      ProcessValue <- "ST_Maintenance_g_u16_5_Times_TiShi_LongDai_Clean"
   Button "按钮_12" at 605,229 size 196x42; TextOff '1小时后提醒 / 1시간후 다시 알림'
      Visibility <- "ST_Maintenance_g_bo_5_Warn_Status_LongDai_Clean"
      on Click: ResetBit("ST_Maintenance_g_bo_5_Warn_Status_LongDai_Clean")
   Button "按钮_13" at 605,282 size 196x42; TextOff '已保养完毕 / 유지보수 이미 완료'; Authorization "User administration"
      Visibility <- "ST_Maintenance_g_bo_5_Warn_Status_LongDai_Clean"
      on Click: ResetBit("ST_Maintenance_g_bo_5_Status_LongDai_Clean")
   TextField "文本域_7" at 61,128 size 812x99; Text '保养时间到,请停机第 次为弓轴滚针 轴承加注黄油 保养时间到,请停机第 次为弓轴滚针 轴承加注黄油 유지보수시간. 기계 스톱. 제 차 보우축 니들 베어링에 그리스를 주입 한다.'
      Visibility <- "ST_Maintenance_g_bo_4_Warn_Status_GongZhou_Bearing"
   IOField "IO Field_90" at 368,129 size 70x28; FormatPattern 999
      Visibility <- "ST_Maintenance_g_bo_4_Warn_Status_GongZhou_Bearing"
      ProcessValue <- "ST_Maintenance_g_u16_4_Times_TiShi_GongZhou_Bearing"
   Button "按钮_10" at 628,129 size 196x42; TextOff '1小时后提醒 / 1시간후 다시 알림'
      Visibility <- "ST_Maintenance_g_bo_4_Warn_Status_GongZhou_Bearing"
      on Click: ResetBit("ST_Maintenance_g_bo_4_Warn_Status_GongZhou_Bearing")
   Button "按钮_11" at 628,182 size 196x42; TextOff '已保养完毕 / 유지보수 이미 완료'; Authorization "User administration"
      Visibility <- "ST_Maintenance_g_bo_4_Warn_Status_GongZhou_Bearing"
      on Click: ResetBit("ST_Maintenance_g_bo_4_Status_GongZhou_Bearing")
   TextField "文本域_9" at 42,238 size 812x100; Text '保养时间到,请停机第 次检查锭子传 动同步带:检查松紧度并适当调整 保养时间到,请停机第 次检查锭子传 动同步带:检查松紧度并适当调整 유지보수시간. 기계 스톱. 제 차 스핀들 전동 타이밍 벨트를 검사 : 조임 정도를 확인 하고 적당하게 조절한다.'
      Visibility <- "ST_Maintenance_g_bo_6_Warn_Status_DingZi_ChuanDong"
   IOField "IO Field_92" at 348,241 size 70x28; FormatPattern 999
      Visibility <- "ST_Maintenance_g_bo_6_Warn_Status_DingZi_ChuanDong"
      ProcessValue <- "ST_Maintenance_g_u16_6_Times_TiShi_DingZi_ChuanDong"
   Button "按钮_14" at 609,240 size 196x42; TextOff '1小时后提醒 / 1시간후 다시 알림'
      Visibility <- "ST_Maintenance_g_bo_6_Warn_Status_DingZi_ChuanDong"
      on Click: ResetBit("ST_Maintenance_g_bo_6_Warn_Status_DingZi_ChuanDong")
   Button "按钮_15" at 609,294 size 196x42; TextOff '已保养完毕 / 유지보수 이미 완료'; Authorization "User administration"
      Visibility <- "ST_Maintenance_g_bo_6_Warn_Status_DingZi_ChuanDong"
      on Click: ResetBit("ST_Maintenance_g_bo_6_Status_DingZi_ChuanDong")
   TextField "文本域_16" at 54,252 size 812x99; Text '保养时间到,请停机第 次清洁控制柜 卫生，用吸风机吸，注意不要用气管吹 保养时间到,请停机第 次清洁控制柜 卫生，用吸风机吸，注意不要用气管吹 유지보수시간. 기계 스톱. 제 차 제어함을 청소 하고 흡입팬으로 흡입한다. 주의할것은 에어 파이프로 불어서는 안된다.'
      Visibility <- "ST_Maintenance_g_bo_7_Warn_Status_ControlBox_Clean"
   IOField "IO Field_98" at 361,254 size 70x28; FormatPattern 999
      Visibility <- "ST_Maintenance_g_bo_7_Warn_Status_ControlBox_Clean"
      ProcessValue <- "ST_Maintenance_g_u16_7_Times_TiShi_ControlBox_Clean"
   Button "按钮_26" at 627,252 size 196x42; TextOff '1小时后提醒 / 1시간후 다시 알림'
      Visibility <- "ST_Maintenance_g_bo_7_Warn_Status_ControlBox_Clean"
      on Click: ResetBit("ST_Maintenance_g_bo_7_Warn_Status_ControlBox_Clean")
   Button "按钮_27" at 627,308 size 196x42; TextOff '已保养完毕 / 유지보수 이미 완료'; Authorization "User administration"
      Visibility <- "ST_Maintenance_g_bo_7_Warn_Status_ControlBox_Clean"
      on Click: ResetBit("ST_Maintenance_g_bo_7_Status_ControlBox_Clean")
   TextField "文本域_13" at 68,268 size 812x99; Text '保养时间到,请停机第 次清洁锭子电 机风扇上的绕毛 保养时间到,请停机第 次清洁锭子电 机风扇上的绕毛 유지보수시간. 기계 스톱. 제 차 스핀들 모터팬 에 감긴 원료 청소한다.'
      Visibility <- "ST_Maintenance_g_bo_8_Warn_Status_DingZi_Fan"
   IOField "IO Field_95" at 373,269 size 70x28; FormatPattern 999
      ProcessValue <- "ST_Maintenance_g_u16_8_Times_TiShi_DingZi_Fan"
      Visibility <- "ST_Maintenance_g_bo_8_Warn_Status_DingZi_Fan"
   Button "按钮_20" at 635,269 size 196x42; TextOff '1小时后提醒 / 1시간후 다시 알림'
      on Click: ResetBit("ST_Maintenance_g_bo_8_Warn_Status_DingZi_Fan")
      Visibility <- "ST_Maintenance_g_bo_8_Warn_Status_DingZi_Fan"
   Button "按钮_21" at 635,324 size 196x41; TextOff '已保养完毕 / 유지보수 이미 완료'; Authorization "User administration"
      on Click: ResetBit("ST_Maintenance_g_bo_8_Status_DingZi_Fan")
      Visibility <- "ST_Maintenance_g_bo_8_Warn_Status_DingZi_Fan"
   Button "按钮_6" at 742,567 size 137x44; TextOff '知道了 / OK'
      on Click: SetTag("ST_HMI_Var_HMI_i16_Dingzi_50102AlarmStatus", 0); ResetBit("ST_HMI_Var_HMI_bo_XiangLing")
      Visibility <- "ST_HMI_Var_HMI_i16_Dingzi_50102AlarmStatus"
   Circle "圆_1" at 782,478 size 60x60
      Visibility <- "ST_HMI_Var_HMI_i16_Dingzi_50102AlarmStatus"
      Appearance <- "ST_HMI_Var_HMI_bo_XiangLing"
   TextField "文本域_5" at 26,442 size 880x170; Text '锭子不转报警！请至报警画面解除报警，然后点击“退 出紧急停止”，点击“启动”开机，或者按正常步骤断电 重启，然后开机 스핀들이 돌아가지 않아 경보알림! 경보알림화면으로 이동하여 경보 해제후 "종료 비상 정지"를 클릭후 "시작"을 클릭하여 가동 하거나 정상적인 순서대로 단전 및 재부팅후 가동한다.'
      Visibility <- "ST_HMI_Var_HMI_i16_Dingzi_50102AlarmStatus"
   Button "按钮_16" at 751,544 size 137x44; TextOff '知道了 / OK'
      on Click: SetTag("ST_HMI_Var_HMI_i16_Dingzi_50102AlarmStatus", 0); ResetBit("ST_HMI_Var_HMI_bo_XiangLing")
      Visibility <- "ST_HMI_Var_HMI_i16_Dingzi_50102AlarmStatus"
   Circle "圆_3" at 791,455 size 60x60
      Visibility <- "ST_HMI_Var_HMI_i16_Dingzi_50102AlarmStatus"
      Appearance <- "ST_HMI_Var_HMI_bo_XiangLing"
   TextField "文本域_11" at 12,427 size 880x170; Text '捻度报警！设置捻度为 ， 实际捻度为 ， 已自动停止，请检查设置画面参数，重新设置总捻度， 检查设置其他参数，使画面上的参数没有红色闪烁，然 后按“启动”，若连续反复出现此报警，请从生头重新 开始 트위스트 경보 알림!설정 트위스트는 이고,실제 트위스트는 이며,이미 자동정지, 설정화면 매개변수를 확인하고,전체 트위스트를 다시 설정하고,기타 매개변수를 확인설정하여 화면의 매개변수에 빨간색이 깜 빡이지 않도록 해야 한다.그다음 "작동"을 누른다. 만약 이 경보가 연속 반 복적으로 나타나면 스레딩부터 다시 시작한다.'
      Visibility <- "ST_HMI_Var_HMI_i16_NianduAlarmStatus"
   IOField "IO Field_43" at 387,432 size 86x32; FormatPattern 9999
      on OnFinishInput: SetBit("ST_Calculation_Var_HMI_bo_Calculation_0_Start"); SetTag("ST_Calculation_Var_g_i16_Calculation_0_3_Select_Status", 1)
      Visibility <- "ST_HMI_Var_HMI_i16_NianduAlarmStatus"
      ProcessValue <- "ST_HMI_Var_HMI_r64NianDu_all"
   IOField "IO Field_3" at 691,432 size 86x32; FormatPattern 9999
      Visibility <- "ST_HMI_Var_HMI_i16_NianduAlarmStatus"
      ProcessValue <- "ST_HMI_Var_HMI_r64Niandu_all_Current"
   Button "按钮_7" at 745,537 size 137x44; TextOff '知道了 / OK'
      on Click: SetTag("ST_HMI_Var_HMI_i16_NianduAlarmStatus", 0); SetBit("ST_Calculation_Var_HMI_bo_Calculation_0_Start"); ResetBit("ST_HMI_Var_HMI_bo_XiangLing")
      Visibility <- "ST_HMI_Var_HMI_i16_NianduAlarmStatus"
   Circle "圆_2" at 785,448 size 60x60
      Visibility <- "ST_HMI_Var_HMI_i16_NianduAlarmStatus"
      Appearance <- "ST_HMI_Var_HMI_bo_XiangLing"

screen "动画" 1280x733, template "模板_2"
   on GenerateScreen: SetTag("变量_100", 9)
   Line "line_3" at 249,441 size 768x20
      Visibility <- "ST_HMI_Var_HMI_r64Axis_1_ZhangLi_Position_JuanRao_real2"
   Line "line_4" at 249,441 size 768x18
      Visibility <- "ST_HMI_Var_HMI_r64Axis_1_ZhangLi_Position_JuanRao_real2"
   Line "line_5" at 251,445 size 766x14
      Visibility <- "ST_HMI_Var_HMI_r64Axis_1_ZhangLi_Position_JuanRao_real2"
   Line "line_6" at 253,449 size 764x10
      Visibility <- "ST_HMI_Var_HMI_r64Axis_1_ZhangLi_Position_JuanRao_real2"
   Line "line_7" at 255,453 size 762x6
      Visibility <- "ST_HMI_Var_HMI_r64Axis_1_ZhangLi_Position_JuanRao_real2"
   Line "line_8" at 255,457 size 762x2
      Visibility <- "ST_HMI_Var_HMI_r64Axis_1_ZhangLi_Position_JuanRao_real2"
   Line "line_12" at 255,459 size 762x6
      Visibility <- "ST_HMI_Var_HMI_r64Axis_1_ZhangLi_Position_JuanRao_real2"
   Line "line_13" at 257,459 size 760x10
      Visibility <- "ST_HMI_Var_HMI_r64Axis_1_ZhangLi_Position_JuanRao_real2"
   Line "line_14" at 257,459 size 760x14
      Visibility <- "ST_HMI_Var_HMI_r64Axis_1_ZhangLi_Position_JuanRao_real2"
   Line "line_27" at 214,457 size 806x20
      Visibility <- "ST_HMI_Var_HMI_r64Axis_1_ZhangLi_Position_JuanRao_real2"
   Line "line_1" at 214,457 size 804x20
      Visibility <- "ST_Main_Var_g_i16_Automatic_Status"
   Group "Group_8" at 262,551 size 1011x176
   Bar "棒图_1" at 177,50 size 20x295; Unit r/min; MinimumValue 0; MaximumValue 10000
      ProcessValue <- "ST_HMI_Var_HMI_r64Axis_DingZi_Velocity_real"
   IOField "IO Field_57" at 166,346 size 62x30; FormatPattern 99999
      ProcessValue <- "ST_HMI_Var_HMI_r64Axis_DingZi_Velocity_real"
   Button "HmiScreenItemData_1" at 1115,95 size 159x60; TextOn '向后 / 後向き / 뒤로'; TextOff '向后 / 後向き / 뒤로'
      on Release: function_efd93a16()
   Rectangle "矩形_3" at 282,425 size 220x80
      DirectMovement <- "ST_HMI_Var_HMI_r64Axis_ZouChe_Position_real2"
   Rectangle "矩形_5" at 486,425 size 214x80
      DirectMovement <- "ST_HMI_Var_HMI_r64Axis_ZouChe_Position_real2"
   Rectangle "矩形_7" at 700,425 size 214x80
      DirectMovement <- "ST_HMI_Var_HMI_r64Axis_ZouChe_Position_real2"
   Rectangle "矩形_8" at 914,425 size 214x80
      DirectMovement <- "ST_HMI_Var_HMI_r64Axis_ZouChe_Position_real2"
   Group "Group_1" at 160,442 size 88x240
   Group "Group_2" at 20,9 size 90x480
   Group "Group_5" at 48,441 size 200x252
   Polyline "折线_1" at 163,442 size 85x231
      Visibility <- "ST_HMI_Var_HMI_r64Axis_ChengXing_Position_real2"
   Polyline "折线_25" at 179,442 size 69x179
      Visibility <- "ST_HMI_Var_HMI_r64Axis_ChengXing_Position_real2"
   Polyline "折线_37" at 197,442 size 51x118
      Visibility <- "ST_HMI_Var_HMI_r64Axis_ChengXing_Position_real2"
   Polyline "折线_45" at 213,442 size 35x57
      Visibility <- "ST_HMI_Var_HMI_r64Axis_ChengXing_Position_real2"
   Polyline "折线_46" at 169,442 size 79x233
      Visibility <- "ST_HMI_Var_HMI_r64Axis_ChengXing_Position_real2"
   Polyline "折线_50" at 179,442 size 69x181
      Visibility <- "ST_HMI_Var_HMI_r64Axis_ChengXing_Position_real2"
   Polyline "折线_51" at 197,442 size 51x122
      Visibility <- "ST_HMI_Var_HMI_r64Axis_ChengXing_Position_real2"
   Polyline "折线_57" at 213,442 size 35x60
      Visibility <- "ST_HMI_Var_HMI_r64Axis_ChengXing_Position_real2"
   Polyline "折线_68" at 169,442 size 79x235
      Visibility <- "ST_HMI_Var_HMI_r64Axis_ChengXing_Position_real2"
   Polyline "折线_71" at 179,442 size 69x184
      Visibility <- "ST_HMI_Var_HMI_r64Axis_ChengXing_Position_real2"
   Polyline "折线_72" at 197,442 size 51x124
      Visibility <- "ST_HMI_Var_HMI_r64Axis_ChengXing_Position_real2"
   Polyline "折线_77" at 213,442 size 35x63
      Visibility <- "ST_HMI_Var_HMI_r64Axis_ChengXing_Position_real2"
   Polyline "折线_78" at 163,442 size 85x237
      Visibility <- "ST_HMI_Var_HMI_r64Axis_ChengXing_Position_real2"
   Polyline "折线_79" at 175,442 size 73x187
      Visibility <- "ST_HMI_Var_HMI_r64Axis_ChengXing_Position_real2"
   Polyline "折线_80" at 191,442 size 57x127
      Visibility <- "ST_HMI_Var_HMI_r64Axis_ChengXing_Position_real2"
   Polyline "折线_81" at 207,442 size 41x66
      Visibility <- "ST_HMI_Var_HMI_r64Axis_ChengXing_Position_real2"
   Polyline "折线_82" at 160,442 size 88x240
      Visibility <- "ST_HMI_Var_HMI_r64Axis_ChengXing_Position_real2"
   Polyline "折线_83" at 207,442 size 41x69
      Visibility <- "ST_HMI_Var_HMI_r64Axis_ChengXing_Position_real2"
   Polyline "折线_84" at 197,442 size 51x131
      Visibility <- "ST_HMI_Var_HMI_r64Axis_ChengXing_Position_real2"
   Polyline "折线_85" at 175,442 size 73x190
      Visibility <- "ST_HMI_Var_HMI_r64Axis_ChengXing_Position_real2"
   Polyline "折线_86" at 175,442 size 73x192
      Visibility <- "ST_HMI_Var_HMI_r64Axis_ChengXing_Position_real2"
   Polyline "折线_87" at 187,442 size 61x133
      Visibility <- "ST_HMI_Var_HMI_r64Axis_ChengXing_Position_real2"
   Polyline "折线_88" at 207,442 size 41x72
      Visibility <- "ST_HMI_Var_HMI_r64Axis_ChengXing_Position_real2"
   Polyline "折线_89" at 179,442 size 69x195
      Visibility <- "ST_HMI_Var_HMI_r64Axis_ChengXing_Position_real2"
   Polyline "折线_90" at 185,442 size 63x136
      Visibility <- "ST_HMI_Var_HMI_r64Axis_ChengXing_Position_real2"
   Polyline "折线_91" at 207,442 size 41x75
      Visibility <- "ST_HMI_Var_HMI_r64Axis_ChengXing_Position_real2"
   Polyline "折线_92" at 175,442 size 73x198
      Visibility <- "ST_HMI_Var_HMI_r64Axis_ChengXing_Position_real2"
   Polyline "折线_93" at 191,442 size 57x140
      Visibility <- "ST_HMI_Var_HMI_r64Axis_ChengXing_Position_real2"
   Polyline "折线_94" at 207,442 size 41x78
      Visibility <- "ST_HMI_Var_HMI_r64Axis_ChengXing_Position_real2"
   Polyline "折线_95" at 175,442 size 73x199
      Visibility <- "ST_HMI_Var_HMI_r64Axis_ChengXing_Position_real2"
   Polyline "折线_96" at 185,442 size 63x143
      Visibility <- "ST_HMI_Var_HMI_r64Axis_ChengXing_Position_real2"
   Polyline "折线_97" at 201,442 size 47x81
      Visibility <- "ST_HMI_Var_HMI_r64Axis_ChengXing_Position_real2"
   Polyline "折线_98" at 175,442 size 73x202
      Visibility <- "ST_HMI_Var_HMI_r64Axis_ChengXing_Position_real2"
   Polyline "折线_99" at 191,442 size 57x146
      Visibility <- "ST_HMI_Var_HMI_r64Axis_ChengXing_Position_real2"
   Polyline "折线_100" at 207,442 size 41x84
      Visibility <- "ST_HMI_Var_HMI_r64Axis_ChengXing_Position_real2"
   Polyline "折线_101" at 167,442 size 81x205
      Visibility <- "ST_HMI_Var_HMI_r64Axis_ChengXing_Position_real2"
   Polyline "折线_102" at 185,442 size 63x149
      Visibility <- "ST_HMI_Var_HMI_r64Axis_ChengXing_Position_real2"
   Polyline "折线_103" at 201,442 size 47x87
      Visibility <- "ST_HMI_Var_HMI_r64Axis_ChengXing_Position_real2"
   Polyline "折线_104" at 169,442 size 79x207
      Visibility <- "ST_HMI_Var_HMI_r64Axis_ChengXing_Position_real2"
   Polyline "折线_105" at 201,442 size 47x91
      Visibility <- "ST_HMI_Var_HMI_r64Axis_ChengXing_Position_real2"
   Polyline "折线_106" at 191,442 size 57x153
      Visibility <- "ST_HMI_Var_HMI_r64Axis_ChengXing_Position_real2"
   Polyline "折线_107" at 169,442 size 79x211
      Visibility <- "ST_HMI_Var_HMI_r64Axis_ChengXing_Position_real2"
   Polyline "折线_108" at 185,442 size 63x156
      Visibility <- "ST_HMI_Var_HMI_r64Axis_ChengXing_Position_real2"
   Polyline "折线_109" at 201,442 size 47x94
      Visibility <- "ST_HMI_Var_HMI_r64Axis_ChengXing_Position_real2"
   Polyline "折线_110" at 169,442 size 79x213
      Visibility <- "ST_HMI_Var_HMI_r64Axis_ChengXing_Position_real2"
   Polyline "折线_111" at 201,442 size 47x96
      Visibility <- "ST_HMI_Var_HMI_r64Axis_ChengXing_Position_real2"
   Polyline "折线_112" at 185,442 size 63x159
      Visibility <- "ST_HMI_Var_HMI_r64Axis_ChengXing_Position_real2"
   Polyline "折线_113" at 170,442 size 78x216
      Visibility <- "ST_HMI_Var_HMI_r64Axis_ChengXing_Position_real2"
   Polyline "折线_114" at 185,442 size 63x161
      Visibility <- "ST_HMI_Var_HMI_r64Axis_ChengXing_Position_real2"
   Polyline "折线_115" at 201,442 size 47x100
      Visibility <- "ST_HMI_Var_HMI_r64Axis_ChengXing_Position_real2"
   Polyline "折线_116" at 179,442 size 69x165
      Visibility <- "ST_HMI_Var_HMI_r64Axis_ChengXing_Position_real2"
   Polyline "折线_117" at 169,442 size 79x219
      Visibility <- "ST_HMI_Var_HMI_r64Axis_ChengXing_Position_real2"
   Polyline "折线_118" at 201,442 size 47x104
      Visibility <- "ST_HMI_Var_HMI_r64Axis_ChengXing_Position_real2"
   Polyline "折线_119" at 169,442 size 79x221
      Visibility <- "ST_HMI_Var_HMI_r64Axis_ChengXing_Position_real2"
   Polyline "折线_120" at 201,442 size 47x106
      Visibility <- "ST_HMI_Var_HMI_r64Axis_ChengXing_Position_real2"
   Polyline "折线_121" at 185,442 size 63x168
      Visibility <- "ST_HMI_Var_HMI_r64Axis_ChengXing_Position_real2"
   Polyline "折线_122" at 169,442 size 79x223
      Visibility <- "ST_HMI_Var_HMI_r64Axis_ChengXing_Position_real2"
   Polyline "折线_123" at 179,442 size 69x170
      Visibility <- "ST_HMI_Var_HMI_r64Axis_ChengXing_Position_real2"
   Polyline "折线_124" at 197,442 size 51x109
      Visibility <- "ST_HMI_Var_HMI_r64Axis_ChengXing_Position_real2"
   Polyline "折线_125" at 165,442 size 83x225
      Visibility <- "ST_HMI_Var_HMI_r64Axis_ChengXing_Position_real2"
   Polyline "折线_126" at 193,442 size 55x112
      Visibility <- "ST_HMI_Var_HMI_r64Axis_ChengXing_Position_real2"
   Polyline "折线_127" at 179,442 size 69x173
      Visibility <- "ST_HMI_Var_HMI_r64Axis_ChengXing_Position_real2"
   Polyline "折线_128" at 169,442 size 79x228
      Visibility <- "ST_HMI_Var_HMI_r64Axis_ChengXing_Position_real2"
   Polyline "折线_129" at 197,442 size 51x115
      Visibility <- "ST_HMI_Var_HMI_r64Axis_ChengXing_Position_real2"
   Polyline "折线_130" at 179,442 size 69x176
      Visibility <- "ST_HMI_Var_HMI_r64Axis_ChengXing_Position_real2"
   Polygon "多边形_195" at 20,131 size 90x323
      Visibility <- "VBS_hengsi_status1"
   Polygon "多边形_196" at 20,229 size 90x225
      Visibility <- "VBS_hengsi_status1"
   Polygon "多边形_264" at 44,338 size 44x116
      Visibility <- "VBS_hengsi_status0"
   Polygon "多边形_265" at 49,350 size 34x104
      Visibility <- "VBS_hengsi_status0"
   Polygon "多边形_198" at 20,124 size 90x330
      Visibility <- "VBS_hengsi_status1"
   Polygon "多边形_199" at 20,223 size 90x231
      Visibility <- "VBS_hengsi_status1"
   Polygon "多边形_266" at 41,329 size 49x124
      Visibility <- "VBS_hengsi_status0"
   Polygon "多边形_201" at 20,120 size 90x334
      Visibility <- "VBS_hengsi_status1"
   Polygon "多边形_202" at 20,219 size 90x235
      Visibility <- "VBS_hengsi_status1"
   Polygon "多边形_267" at 38,319 size 54x135
      Visibility <- "VBS_hengsi_status0"
   Polygon "多边形_204" at 20,117 size 90x337
      Visibility <- "VBS_hengsi_status1"
   Polygon "多边形_205" at 20,213 size 90x241
      Visibility <- "VBS_hengsi_status1"
   Polygon "多边形_268" at 36,311 size 58x143
      Visibility <- "VBS_hengsi_status0"
   Polygon "多边形_207" at 20,113 size 90x341
      Visibility <- "VBS_hengsi_status1"
   Polygon "多边形_208" at 20,210 size 90x243
      Visibility <- "VBS_hengsi_status1"
   Polygon "多边形_269" at 35,306 size 60x148
      Visibility <- "VBS_hengsi_status0"
   Polygon "多边形_210" at 20,107 size 90x347
      Visibility <- "VBS_hengsi_status0"
   Polygon "多边形_211" at 20,206 size 90x248
      Visibility <- "VBS_hengsi_status1"
   Polygon "多边形_270" at 35,298 size 60x156
      Visibility <- "VBS_hengsi_status0"
   Polygon "多边形_213" at 20,103 size 90x351
      Visibility <- "VBS_hengsi_status1"
   Polygon "多边形_214" at 20,202 size 90x252
      Visibility <- "VBS_hengsi_status1"
   Polygon "多边形_271" at 34,292 size 63x162
      Visibility <- "VBS_hengsi_status0"
   Polygon "多边形_216" at 20,97 size 90x357
      Visibility <- "VBS_hengsi_status1"
   Polygon "多边形_217" at 20,196 size 90x258
      Visibility <- "VBS_hengsi_status1"
   Polygon "多边形_272" at 34,288 size 63x166
      Visibility <- "VBS_hengsi_status0"
   Polygon "多边形_219" at 20,93 size 90x361
      Visibility <- "VBS_hengsi_status1"
   Polygon "多边形_220" at 20,192 size 90x262
      Visibility <- "VBS_hengsi_status1"
   Polygon "多边形_273" at 32,285 size 66x169
      Visibility <- "VBS_hengsi_status0"
   Polygon "多边形_222" at 20,90 size 90x364
      Visibility <- "VBS_hengsi_status1"
   Polygon "多边形_223" at 20,189 size 90x265
      Visibility <- "VBS_hengsi_status1"
   Polygon "多边形_274" at 32,283 size 66x171
      Visibility <- "VBS_hengsi_status0"
   Polygon "多边形_225" at 20,86 size 90x368
      Visibility <- "VBS_hengsi_status1"
   Polygon "多边形_226" at 20,185 size 90x269
      Visibility <- "VBS_hengsi_status1"
   Polygon "多边形_275" at 31,279 size 68x175
      Visibility <- "VBS_hengsi_status0"
   Polygon "多边形_228" at 20,80 size 90x374
      Visibility <- "VBS_hengsi_status1"
   Polygon "多边形_229" at 20,179 size 90x275
      Visibility <- "VBS_hengsi_status1"
   Polygon "多边形_276" at 31,275 size 68x179
      Visibility <- "VBS_hengsi_status0"
   Polygon "多边形_231" at 20,76 size 90x378
      Visibility <- "VBS_hengsi_status1"
   Polygon "多边形_232" at 20,175 size 90x279
      Visibility <- "VBS_hengsi_status1"
   Polygon "多边形_277" at 29,271 size 70x183
      Visibility <- "VBS_hengsi_status0"
   Polygon "多边形_234" at 20,70 size 90x384
      Visibility <- "VBS_hengsi_status1"
   Polygon "多边形_235" at 20,169 size 90x285
      Visibility <- "VBS_hengsi_status1"
   Polygon "多边形_278" at 27,271 size 74x183
      Visibility <- "VBS_hengsi_status0"
   Polygon "多边形_237" at 20,69 size 90x385
      Visibility <- "VBS_hengsi_status1"
   Polygon "多边形_238" at 20,165 size 90x289
      Visibility <- "VBS_hengsi_status1"
   Polygon "多边形_279" at 27,267 size 74x187
      Visibility <- "VBS_hengsi_status0"
   Polygon "多边形_240" at 20,63 size 90x391
      Visibility <- "VBS_hengsi_status1"
   Polygon "多边形_241" at 20,162 size 90x292
      Visibility <- "VBS_hengsi_status1"
   Polygon "多边形_280" at 26,263 size 77x191
      Visibility <- "VBS_hengsi_status0"
   Polygon "多边形_243" at 20,59 size 90x395
      Visibility <- "VBS_hengsi_status1"
   Polygon "多边形_244" at 20,158 size 90x296
      Visibility <- "VBS_hengsi_status1"
   Polygon "多边形_281" at 26,261 size 77x193
      Visibility <- "VBS_hengsi_status0"
   Polygon "多边形_246" at 20,53 size 90x401
      Visibility <- "VBS_hengsi_status1"
   Polygon "多边形_247" at 20,152 size 90x302
      Visibility <- "VBS_hengsi_status1"
   Polygon "多边形_282" at 25,258 size 79x196
      Visibility <- "VBS_hengsi_status0"
   Polygon "多边形_249" at 20,49 size 90x405
      Visibility <- "VBS_hengsi_status1"
   Polygon "多边形_250" at 20,148 size 90x306
      Visibility <- "VBS_hengsi_status1"
   Polygon "多边形_283" at 25,254 size 79x200
      Visibility <- "VBS_hengsi_status0"
   Polygon "多边形_252" at 20,45 size 90x409
      Visibility <- "VBS_hengsi_status1"
   Polygon "多边形_253" at 20,142 size 90x312
      Visibility <- "VBS_hengsi_status1"
   Polygon "多边形_284" at 23,250 size 83x204
      Visibility <- "VBS_hengsi_status0"
   Polygon "多边形_255" at 20,42 size 90x412
      Visibility <- "VBS_hengsi_status1"
   Polygon "多边形_256" at 20,141 size 90x313
      Visibility <- "VBS_hengsi_status1"
   Polygon "多边形_285" at 23,246 size 83x208
      Visibility <- "VBS_hengsi_status0"
   Polygon "多边形_258" at 20,135 size 90x319
      Visibility <- "VBS_hengsi_status1"
   Polygon "多边形_286" at 22,242 size 85x212
      Visibility <- "VBS_hengsi_status0"
   Polygon "多边形_287" at 22,238 size 85x216
      Visibility <- "VBS_hengsi_status0"
   Polygon "多边形_288" at 20,237 size 88x217
      Visibility <- "VBS_hengsi_status0"
   Polygon "多边形_289" at 20,231 size 90x223
      Visibility <- "VBS_hengsi_status0"
   Group "Group_3" at 48,441 size 200x252
   Group "Group_4" at 48,441 size 200x252
   Line "线_1" at 68,549 size 180x9
      Visibility <- "ST_HMI_Var_HMI_r64Axis_ChengXing_Position_real2"
   Line "线_2" at 68,549 size 166x68
      Visibility <- "ST_HMI_Var_HMI_r64Axis_ChengXing_Position_real2"
   Line "线_136#mig1_2" at 68,549 size 132x120
      Visibility <- "ST_HMI_Var_HMI_r64Axis_ChengXing_Position_real2"
   Line "线_3" at 68,443 size 144x106
      Visibility <- "ST_HMI_Var_HMI_r64Axis_ChengXing_Position_real2"
   Line "线_4" at 68,497 size 172x52
      Visibility <- "ST_HMI_Var_HMI_r64Axis_ChengXing_Position_real2"
   Line "线_11#mig1_2" at 68,441 size 143x108
      Visibility <- "ST_HMI_Var_HMI_r64Axis_ChengXing_Position_real2"
   Line "线_5" at 68,501 size 173x48
      Visibility <- "ST_HMI_Var_HMI_r64Axis_ChengXing_Position_real2"
   Line "线_6" at 68,549 size 129x122
      Visibility <- "ST_HMI_Var_HMI_r64Axis_ChengXing_Position_real2"
   Line "线_157" at 68,446 size 146x103
      Visibility <- "ST_HMI_Var_HMI_r64Axis_ChengXing_Position_real2"
   Line "线_115#mig1_2" at 68,549 size 179x13
      Visibility <- "ST_HMI_Var_HMI_r64Axis_ChengXing_Position_real2"
   Line "线_7" at 68,549 size 165x71
      Visibility <- "ST_HMI_Var_HMI_r64Axis_ChengXing_Position_real2"
   Line "线_159" at 68,549 size 179x15
      Visibility <- "ST_HMI_Var_HMI_r64Axis_ChengXing_Position_real2"
   Line "线_8" at 68,549 size 163x74
      Visibility <- "ST_HMI_Var_HMI_r64Axis_ChengXing_Position_real2"
   Line "线_9" at 68,549 size 127x124
      Visibility <- "ST_HMI_Var_HMI_r64Axis_ChengXing_Position_real2"
   Line "线_13#mig1_2" at 68,448 size 147x101
      Visibility <- "ST_HMI_Var_HMI_r64Axis_ChengXing_Position_real2"
   Line "线_14" at 68,503 size 174x46
      Visibility <- "ST_HMI_Var_HMI_r64Axis_ChengXing_Position_real2"
   Line "线_22" at 68,549 size 179x18
      Visibility <- "ST_HMI_Var_HMI_r64Axis_ChengXing_Position_real2"
   Line "线_24" at 68,549 size 162x77
      Visibility <- "ST_HMI_Var_HMI_r64Axis_ChengXing_Position_real2"
   Line "线_25" at 68,549 size 125x126
      Visibility <- "ST_HMI_Var_HMI_r64Axis_ChengXing_Position_real2"
   Line "线_124#mig1_2" at 68,451 size 149x98
      Visibility <- "ST_HMI_Var_HMI_r64Axis_ChengXing_Position_real2"
   Line "线_27" at 68,507 size 175x42
      Visibility <- "ST_HMI_Var_HMI_r64Axis_ChengXing_Position_real2"
   Line "线_195" at 68,549 size 179x21
      Visibility <- "ST_HMI_Var_HMI_r64Axis_ChengXing_Position_real2"
   Line "线_196" at 68,549 size 161x80
      Visibility <- "ST_HMI_Var_HMI_r64Axis_ChengXing_Position_real2"
   Line "线_197" at 68,549 size 122x129
      Visibility <- "ST_HMI_Var_HMI_r64Axis_ChengXing_Position_real2"
   Line "线_198" at 68,454 size 151x95
      Visibility <- "ST_HMI_Var_HMI_r64Axis_ChengXing_Position_real2"
   Line "线_199" at 68,510 size 175x39
      Visibility <- "ST_HMI_Var_HMI_r64Axis_ChengXing_Position_real2"
   Line "线_200" at 68,549 size 178x24
      Visibility <- "ST_HMI_Var_HMI_r64Axis_ChengXing_Position_real2"
   Line "线_201" at 68,549 size 159x82
      Visibility <- "ST_HMI_Var_HMI_r64Axis_ChengXing_Position_real2"
   Line "线_202" at 68,549 size 120x131
      Visibility <- "ST_HMI_Var_HMI_r64Axis_ChengXing_Position_real2"
   Line "线_254" at 68,456 size 153x93
      Visibility <- "ST_HMI_Var_HMI_r64Axis_ChengXing_Position_real2"
   Line "线_255" at 68,513 size 176x36
      Visibility <- "ST_HMI_Var_HMI_r64Axis_ChengXing_Position_real2"
   Line "线_256" at 68,549 size 178x27
      Visibility <- "ST_HMI_Var_HMI_r64Axis_ChengXing_Position_real2"
   Line "线_257" at 68,549 size 157x85
      Visibility <- "ST_HMI_Var_HMI_r64Axis_ChengXing_Position_real2"
   Line "线_277" at 68,549 size 118x133
      Visibility <- "ST_HMI_Var_HMI_r64Axis_ChengXing_Position_real2"
   Line "线_278" at 68,459 size 154x90
      Visibility <- "ST_HMI_Var_HMI_r64Axis_ChengXing_Position_real2"
   Line "线_279" at 68,516 size 177x33
      Visibility <- "ST_HMI_Var_HMI_r64Axis_ChengXing_Position_real2"
   Line "线_280" at 68,549 size 177x31
      Visibility <- "ST_HMI_Var_HMI_r64Axis_ChengXing_Position_real2"
   Line "线_281" at 68,549 size 156x88
      Visibility <- "ST_HMI_Var_HMI_r64Axis_ChengXing_Position_real2"
   Line "线_282" at 68,549 size 116x135
      Visibility <- "ST_HMI_Var_HMI_r64Axis_ChengXing_Position_real2"
   Line "线_283" at 68,462 size 156x87
      Visibility <- "ST_HMI_Var_HMI_r64Axis_ChengXing_Position_real2"
   Line "线_125#mig1_2" at 68,518 size 177x31
      Visibility <- "ST_HMI_Var_HMI_r64Axis_ChengXing_Position_real2"
   Line "线_284" at 68,549 size 177x33
      Visibility <- "ST_HMI_Var_HMI_r64Axis_ChengXing_Position_real2"
   Line "线_285" at 68,549 size 154x90
      Visibility <- "ST_HMI_Var_HMI_r64Axis_ChengXing_Position_real2"
   Line "线_286" at 68,549 size 113x137
      Visibility <- "ST_HMI_Var_HMI_r64Axis_ChengXing_Position_real2"
   Line "线_287" at 68,464 size 157x85
      Visibility <- "ST_HMI_Var_HMI_r64Axis_ChengXing_Position_real2"
   Line "线_288" at 68,521 size 178x28
      Visibility <- "ST_HMI_Var_HMI_r64Axis_ChengXing_Position_real2"
   Line "线_289" at 68,549 size 176x37
      Visibility <- "ST_HMI_Var_HMI_r64Axis_ChengXing_Position_real2"
   Line "线_290" at 68,549 size 153x93
      Visibility <- "ST_HMI_Var_HMI_r64Axis_ChengXing_Position_real2"
   Line "线_291" at 68,549 size 111x139
      Visibility <- "ST_HMI_Var_HMI_r64Axis_ChengXing_Position_real2"
   Line "线_292" at 68,466 size 159x83
      Visibility <- "ST_HMI_Var_HMI_r64Axis_ChengXing_Position_real2"
   Line "线_293" at 68,524 size 179x25
      Visibility <- "ST_HMI_Var_HMI_r64Axis_ChengXing_Position_real2"
   Line "线_294" at 68,549 size 175x39
      Visibility <- "ST_HMI_Var_HMI_r64Axis_ChengXing_Position_real2"
   Line "线_295" at 68,549 size 151x96
      Visibility <- "ST_HMI_Var_HMI_r64Axis_ChengXing_Position_real2"
   Line "线_315" at 68,549 size 108x141
      Visibility <- "ST_HMI_Var_HMI_r64Axis_ChengXing_Position_real2"
   Line "线_316" at 68,469 size 161x80
      Visibility <- "ST_HMI_Var_HMI_r64Axis_ChengXing_Position_real2"
   Line "线_130#mig1_2" at 68,527 size 179x22
      Visibility <- "ST_HMI_Var_HMI_r64Axis_ChengXing_Position_real2"
   Line "线_317" at 68,549 size 106x143
      Visibility <- "ST_HMI_Var_HMI_r64Axis_ChengXing_Position_real2"
   Line "线_97#mig1_2" at 68,471 size 162x78
      Visibility <- "ST_HMI_Var_HMI_r64Axis_ChengXing_Position_real2"
   Line "线_129#mig1_2" at 68,530 size 179x19
      Visibility <- "ST_HMI_Var_HMI_r64Axis_ChengXing_Position_real2"
   Line "线_318" at 68,549 size 175x43
      Visibility <- "ST_HMI_Var_HMI_r64Axis_ChengXing_Position_real2"
   Line "线_319" at 68,549 size 149x98
      Visibility <- "ST_HMI_Var_HMI_r64Axis_ChengXing_Position_real2"
   Line "线_320" at 68,549 size 103x144
      Visibility <- "ST_HMI_Var_HMI_r64Axis_ChengXing_Position_real2"
   Line "线_321" at 68,474 size 163x75
      Visibility <- "ST_HMI_Var_HMI_r64Axis_ChengXing_Position_real2"
   Line "线_128#mig1_2" at 68,534 size 179x15
      Visibility <- "ST_HMI_Var_HMI_r64Axis_ChengXing_Position_real2"
   Line "线_322" at 68,549 size 174x46
      Visibility <- "ST_HMI_Var_HMI_r64Axis_ChengXing_Position_real2"
   Line "线_323" at 68,549 size 147x101
      Visibility <- "ST_HMI_Var_HMI_r64Axis_ChengXing_Position_real2"
   Line "线_324" at 68,477 size 165x72
      Visibility <- "ST_HMI_Var_HMI_r64Axis_ChengXing_Position_real2"
   Line "线_131#mig1_2" at 68,536 size 179x13
      Visibility <- "ST_HMI_Var_HMI_r64Axis_ChengXing_Position_real2"
   Line "线_325" at 68,549 size 173x49
      Visibility <- "ST_HMI_Var_HMI_r64Axis_ChengXing_Position_real2"
   Line "线_326" at 68,549 size 146x104
      Visibility <- "ST_HMI_Var_HMI_r64Axis_ChengXing_Position_real2"
   Line "线_114#mig1_2" at 68,480 size 166x69
      Visibility <- "ST_HMI_Var_HMI_r64Axis_ChengXing_Position_real2"
   Line "线_327" at 68,540 size 180x9
      Visibility <- "ST_HMI_Var_HMI_r64Axis_ChengXing_Position_real2"
   Line "线_328" at 68,549 size 172x52
      Visibility <- "ST_HMI_Var_HMI_r64Axis_ChengXing_Position_real2"
   Line "线_329" at 68,549 size 144x106
      Visibility <- "ST_HMI_Var_HMI_r64Axis_ChengXing_Position_real2"
   Line "线_120#mig1_2" at 68,483 size 167x66
      Visibility <- "ST_HMI_Var_HMI_r64Axis_ChengXing_Position_real2"
   Line "线_330" at 68,543 size 180x6
      Visibility <- "ST_HMI_Var_HMI_r64Axis_ChengXing_Position_real2"
   Line "线_331" at 68,549 size 171x55
      Visibility <- "ST_HMI_Var_HMI_r64Axis_ChengXing_Position_real2"
   Line "线_332" at 68,549 size 142x109
      Visibility <- "ST_HMI_Var_HMI_r64Axis_ChengXing_Position_real2"
   Line "线_333" at 68,486 size 168x63
      Visibility <- "ST_HMI_Var_HMI_r64Axis_ChengXing_Position_real2"
   Line "线_150#mig1_2" at 68,546 size 180x3
      Visibility <- "ST_HMI_Var_HMI_r64Axis_ChengXing_Position_real2"
   Line "线_334" at 68,549 size 170x58
      Visibility <- "ST_HMI_Var_HMI_r64Axis_ChengXing_Position_real2"
   Line "线_335" at 68,549 size 140x111
      Visibility <- "ST_HMI_Var_HMI_r64Axis_ChengXing_Position_real2"
   Line "线_336" at 68,489 size 169x60
      Visibility <- "ST_HMI_Var_HMI_r64Axis_ChengXing_Position_real2"
   Line "线_147#mig1_2" at 68,549 size 180x0
      Visibility <- "ST_HMI_Var_HMI_r64Axis_ChengXing_Position_real2"
   Line "线_337" at 68,549 size 169x61
      Visibility <- "ST_HMI_Var_HMI_r64Axis_ChengXing_Position_real2"
   Line "线_338" at 68,549 size 138x114
      Visibility <- "ST_HMI_Var_HMI_r64Axis_ChengXing_Position_real2"
   Line "线_339" at 68,491 size 170x58
      Visibility <- "ST_HMI_Var_HMI_r64Axis_ChengXing_Position_real2"
   Line "线_340" at 68,549 size 180x3
      Visibility <- "ST_HMI_Var_HMI_r64Axis_ChengXing_Position_real2"
   Line "线_341" at 68,549 size 168x63
      Visibility <- "ST_HMI_Var_HMI_r64Axis_ChengXing_Position_real2"
   Line "线_342" at 68,549 size 167x67
      Visibility <- "ST_HMI_Var_HMI_r64Axis_ChengXing_Position_real2"
   Line "线_343" at 68,549 size 136x116
      Visibility <- "ST_HMI_Var_HMI_r64Axis_ChengXing_Position_real2"
   Line "线_344" at 68,549 size 134x118
      Visibility <- "ST_HMI_Var_HMI_r64Axis_ChengXing_Position_real2"
   Line "线_345" at 68,495 size 171x54